         i18 : Int;
         i19 : Int;
         i20 : Int;
         i21 : Int;
      END_STRUCT;
      STC_tMngSysReg : Struct   // Managment system register
         tST : Struct
            xWrite_Request : Bool;
            xDone : Bool;
            xBusy : Bool;
            xError : Bool;
            xSpare4 : Bool;
            xSpare5 : Bool;
            xSpare6 : Bool;
            xSpare7 : Bool;
            ID : Hw_Io;
            dINDEX : DInt;
            uiLEN : UInt;
            dwSTATUS : DWord;
            iSpare : Int;
         END_STRUCT;
         tDATA : Struct
            wRequest_refere_RequestID : Word := W#16#102;   // (Request_referece=01 Alwais=01 )*(RequestID=02 Change Param)
            wAxis_NoOfParameters : Word := W#16#101;   // (Axis=Num.Object)(NoOfParameters=Num of parameter to change)
            wAttribute_NoOfElements : Word := W#16#1001;   // (Attribute=10 Alwais=10)(NoOfParameters=Num of subparameter to Write)
            iParameter_number : Int := 2599;   // Parameter_number=Number of the parameter
            wSubindex : Word;   // Subindex
            wFormat_NoOfValue : Word := W#16#4301;   // (Format_NoOfValue=Format 42=Word 43=Dword)(Num. of value to transfer)
            dwRegisterValue : DWord := DW#16#1;   // Register value
         END_STRUCT;
      END_STRUCT;
      STC_tWriteRecord : WRREC;
      STC_tPZD_OpCLLoop : Struct   // Motor module open/close loop telegram 1
         tR : Struct   // READ
            tZSW1 : Struct   // R2089[0].STATUS WORD 1
               x8 : Bool;   // Speed setp-act val deviation in tollerance
               x9 : Bool;   // Control request
               x10 : Bool;   // F or n comparision value reached or exceeded
               x11 : Bool;   // Tourque limit reached
               x12 : Bool;   // Open holding brake
               x13 : Bool;   // Alarm motor overtemperature
               x14 : Bool;   // n_act>=0
               x15 : Bool;   // Alarm power unit thermal overload
               x0 : Bool;   // Ready for switch on
               x1 : Bool;   // Ready
               x2 : Bool;   // Operation enabled
               x3 : Bool;   // Fault present
               x4 : Bool;   // OFF2
               x5 : Bool;   // OFF3
               x6 : Bool;   // Switching on inhibited active
               x7 : Bool;   // Alarm present
            END_STRUCT;
            iNIST_A : Int;   // R63.Actual speed value
            iFAULT_CODE : Int;   // R2131.Actual fault code
            iWARN_CODE : Int;   // R2132.Actual alarm code
            iUserData1 : Int;
            iUserData2 : Int;
         END_STRUCT;
         tW : Struct   // WRITE
            tSTW1 : Struct   // CONTROL WORD 1
               x8 : Bool;   // Reserved
               x9 : Bool;   // P1122[0].Bypass ramp-function generator
               x10 : Bool;   // P854[0].Control by PLC
               x11 : Bool;   // P1113[0].Setpoint inversion
               x12 : Bool;   // Reserved
               x13 : Bool;   // P1035[0].Motorized potentiometer setpoint raise
               x14 : Bool;   // P1036[0].Motorized potentiometer setpoint lower
               x15 : Bool;   // P855[0] Brake release
               x0 : Bool;   // P840[0].ON/OFF
               x1 : Bool;   // P844[0].OFF2
               x2 : Bool;   // P848[0].OFF3
               x3 : Bool;   // P852[0].Enable operation
               x4 : Bool;   // P1140[0].Enable ramp function generator
               x5 : Bool;   // P1141[0].Continue ramp function generator
               x6 : Bool;   // P1142[0].Enable setpoint
               x7 : Bool;   // P2103[0].Acknowledge faults
            END_STRUCT;
            iNSOLL_A : Int;   // P1070[0].Main set point
            iACC : Int;   // P1138[0].Acceleration ramp % [0-16384]
            iDEC : Int;   // P1139[0].Deceleration ramp % [0-16384]
            iExtRef : Int;   // P1076[0].External reference scaling % [0-16384]
            iUserData2 : Int;
         END_STRUCT;
      END_STRUCT;
   END_VAR
   VAR_TEMP
      TMP_dOldValue_AR1 : DInt;
      TMP_dOldValue_AR2 : DInt;
      TMP_x : Bool;
      TMP_i : Int;
      TMP_d : DInt;
      TMP_r : Real;
      TMP_a : ANY;
      TMP_dZero : DInt;
      TMP_xAlwaysON : Bool;
      TMP_rActualSpeed : Real;
      TMP_iAddressLength : Int;
      TMP_dActualPosMin_dmm : DInt;   // Actual position minimum tollerance [mm/10]
      TMP_dActualPosMax_dmm : DInt;   // Actual position maximum tollerance [mm/10]
      TMP_iRetVal : Int;
   END_VAR
BEGIN

REGION Network 1 (STL): Save AR1 & AR2 value
   //    TAR1
   //    T     #TMP_dOldValue_AR1
   //    TAR2
   //    T     #TMP_dOldValue_AR2
END_REGION

REGION Network 2: #####_COSTANTS_#####
END_REGION

REGION Network 3 (STL): Initializing
         SET;
         S     #TMP_xAlwaysON;

         L     DINT#0;
         T     #TMP_dZero;


         CALL  FILL
         ( BVAL    := #TMP_dZero,
           RET_VAL := #TMP_iRetVal,
           BLK     := #STC_tPZD_OpCLLoop.tR
         );

         CALL  FILL
         ( BVAL    := #TMP_dZero,
           RET_VAL := #TMP_iRetVal,
           BLK     := #STC_tMngSysReg
         );
END_REGION

REGION Network 4: #####_MOTOR_MODULE_#####
END_REGION

REGION Network 5 (STL): Check system data coerence
         L     #STC_tSYS_DATA.iIOAddress_MM;
         L     0;
         <I;
         L     10;
         JC    Err;

         L     #STC_tSYS_DATA.dMaxSpeed_rpm;
         L     DINT#0;
         <=D;
         L     11;
         JC    Err;

         L     #STC_tSYS_DATA.rK_rpm_mmMin;
         L     0.0;
         <=R;
         L     12;
         JC    Err;

         L     #STC_tSYS_DATA.rK_mmMin_Rpm;
         L     0.0;
         <=R;
         L     13;
         JC    Err;

         L     #STC_tSYS_DATA.rMaxAcc_s;
         L     0.0;
         <=R;
         L     14;
         JC    Err;

         L     #STC_tSYS_DATA.rMaxDec_s;
         L     0.0;
         <=R;
         L     15;
         JC    Err;

         L     6;
         T     #TMP_iAddressLength;

   //Compute destination position
         L;
         LAR1;
   //byte 1 = 10h (FIXED for S7)
         L     B#16#10;
         T     B[AR1, P#0.0];
   //byte 2 = data type
         L     B#16#4;  //4 = word
         T     B[AR1, P#1.0];
   //byte 3 & 4 = number of element
         L     #TMP_iAddressLength;  //Production data
         T     W[AR1, P#2.0];
   //byte 5 & 6 = number of DB
         L     0;  //DB production data
         T     W[AR1, P#4.0];
   //byte 7 = memory area
         L     B#16#81;  //81h = I (Input)
         T     B[AR1, P#6.0];
   //byte 8 & 9 = address. Bit 0,1,2 of tenth byte is bit offset
   //byte 7 = address (high). Valid value = 0-7. Bit 3,4,5,6,7 always 0

         L     #STC_tSYS_DATA.iIOAddress_MM;  //Item size
         SLW   3;
         T     W[AR1, P#8.0];
         SRD   16;
         AW    16#0007;
         T     B[AR1, P#7.0];
END_REGION

REGION Network 6: ########################_OPEN_CLOSE_LOOP_#######################
END_REGION

REGION Network 7: #####_MATCH_#####
END_REGION

REGION Network 8 (STL): Input copy
         CALL  BLKMOV
         ( SRCBLK  := #TMP_a,
           RET_VAL := #TMP_iRetVal,
           DSTBLK  := #STC_tPZD_OpCLLoop.tR
         );
END_REGION

REGION Network 9: Status signals
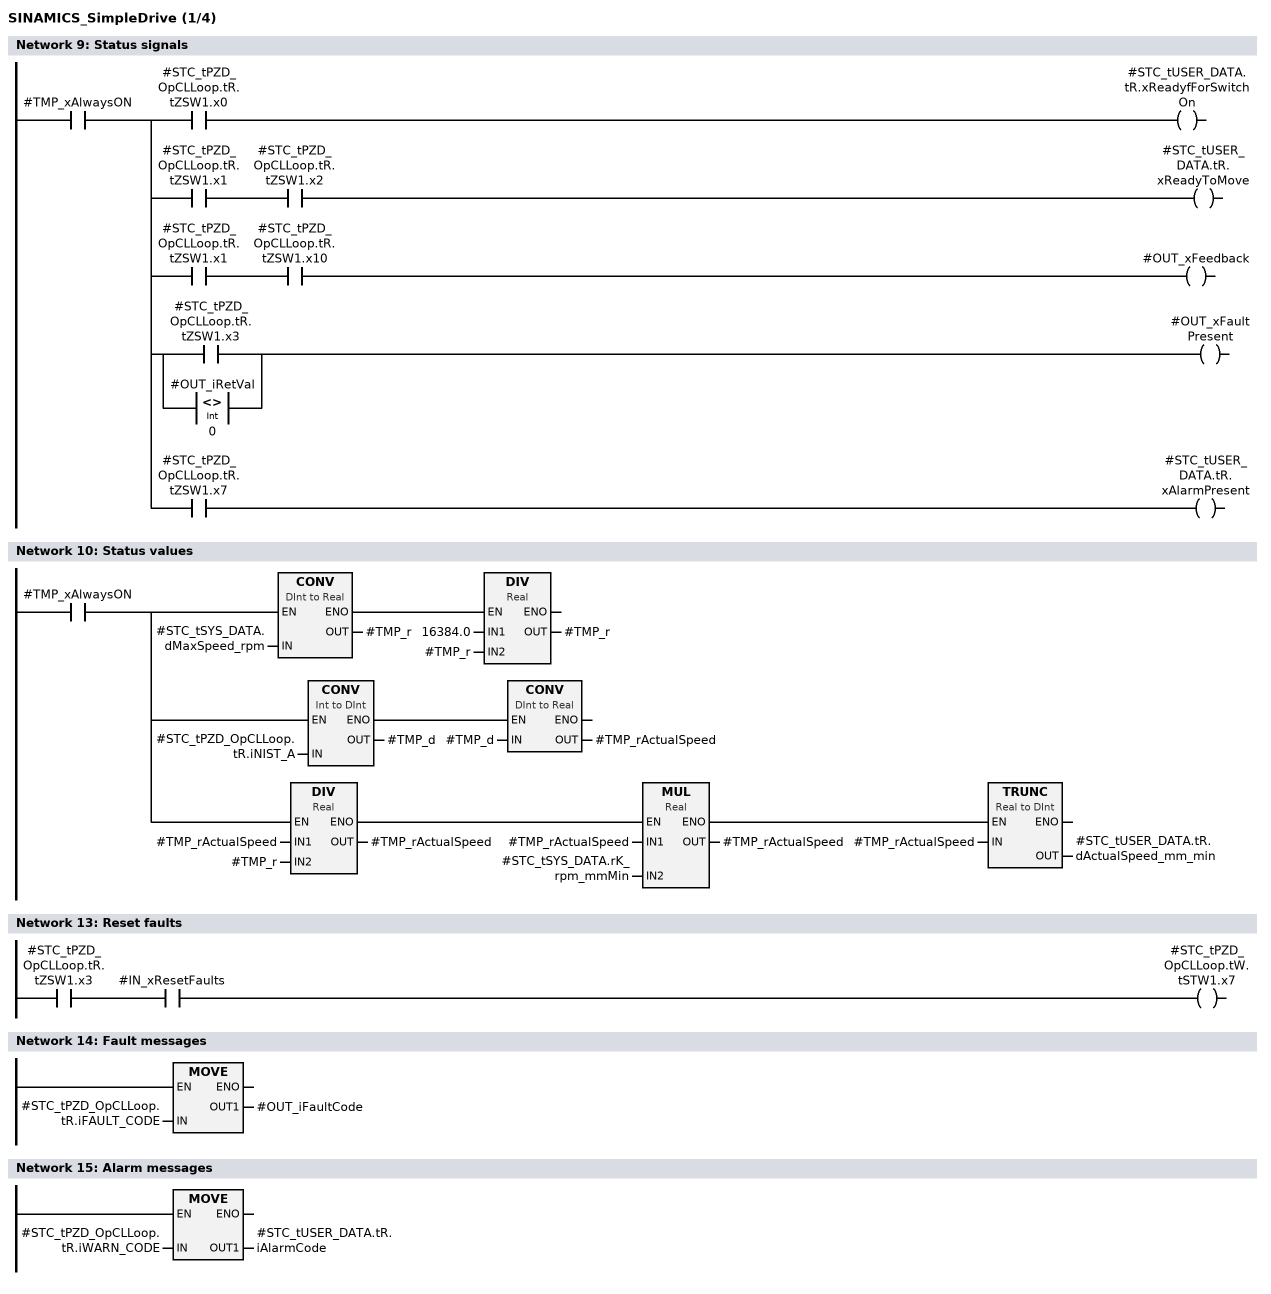
   RUNG wire#powerrail
      Contact( #TMP_xAlwaysON )
      wire#w1
      Contact( #STC_tPZD_OpCLLoop.tR.tZSW1.x0 )
      Coil( #STC_tUSER_DATA.tR.xReadyfForSwitchOn )
   END_RUNG
   RUNG wire#w1
      Contact( #STC_tPZD_OpCLLoop.tR.tZSW1.x1 )
      Contact( #STC_tPZD_OpCLLoop.tR.tZSW1.x2 )
      Coil( #STC_tUSER_DATA.tR.xReadyToMove )
   END_RUNG
   RUNG wire#w1
      Contact( #STC_tPZD_OpCLLoop.tR.tZSW1.x1 )
      Contact( #STC_tPZD_OpCLLoop.tR.tZSW1.x10 )
      Coil( #OUT_xFeedback )
   END_RUNG
   RUNG wire#w1
      Contact( #STC_tPZD_OpCLLoop.tR.tZSW1.x3 )
      wire#w2
      Coil( #OUT_xFaultPresent )
   END_RUNG
   RUNG wire#w1
      { S7_Templates := "SrcType := Int" } NE_Contact(in1 := #OUT_iRetVal, in2 := 0)
   END_RUNG wire#w2
   RUNG wire#w1
      Contact( #STC_tPZD_OpCLLoop.tR.tZSW1.x7 )
      Coil( #STC_tUSER_DATA.tR.xAlarmPresent )
   END_RUNG
   // the same network as SCL:
   #STC_tUSER_DATA.tR.xReadyfForSwitchOn := #TMP_xAlwaysON AND #STC_tPZD_OpCLLoop.tR.tZSW1.x0;
   #STC_tUSER_DATA.tR.xReadyToMove := #TMP_xAlwaysON AND #STC_tPZD_OpCLLoop.tR.tZSW1.x1 AND #STC_tPZD_OpCLLoop.tR.tZSW1.x2;
   #OUT_xFeedback := #TMP_xAlwaysON AND #STC_tPZD_OpCLLoop.tR.tZSW1.x1 AND #STC_tPZD_OpCLLoop.tR.tZSW1.x10;
   #OUT_xFaultPresent := #TMP_xAlwaysON AND (#STC_tPZD_OpCLLoop.tR.tZSW1.x3 OR (#OUT_iRetVal <> 0));
   #STC_tUSER_DATA.tR.xAlarmPresent := #TMP_xAlwaysON AND #STC_tPZD_OpCLLoop.tR.tZSW1.x7;
END_REGION

REGION Network 10: Status values
   RUNG wire#powerrail
      Contact( #TMP_xAlwaysON )
      wire#w1
      { S7_Templates := "[SrcType := DInt, DestType := Real]"; S7_GenerateENO := "TRUE" } Convert(in := #STC_tSYS_DATA.dMaxSpeed_rpm, out => #TMP_r)
      { S7_Templates := "SrcType := Real"; S7_GenerateENO := "TRUE" } Div(in1 := 16384.0, in2 := #TMP_r, out => #TMP_r)
   END_RUNG
   RUNG wire#w1
      { S7_Templates := "[SrcType := Int, DestType := DInt]"; S7_GenerateENO := "TRUE" } Convert(in := #STC_tPZD_OpCLLoop.tR.iNIST_A, out => #TMP_d)
      { S7_Templates := "[SrcType := DInt, DestType := Real]"; S7_GenerateENO := "TRUE" } Convert(in := #TMP_d, out => #TMP_rActualSpeed)
   END_RUNG
   RUNG wire#w1
      { S7_Templates := "SrcType := Real"; S7_GenerateENO := "TRUE" } Div(in1 := #TMP_rActualSpeed, in2 := #TMP_r, out => #TMP_rActualSpeed)
      { S7_Templates := "SrcType := Real"; S7_GenerateENO := "TRUE" } Mul(in1 := #TMP_rActualSpeed, in2 := #STC_tSYS_DATA.rK_rpm_mmMin, out => #TMP_rActualSpeed)
      { S7_Templates := "[SrcType := Real, DestType := DInt]"; S7_GenerateENO := "TRUE" } Trunc(in := #TMP_rActualSpeed, out => #STC_tUSER_DATA.tR.dActualSpeed_mm_min)
   END_RUNG
   // the same network as SCL:
   // ENO of a box is taken as its EN; it also drops when the box reports an error
   IF #TMP_xAlwaysON THEN
       #TMP_r := DINT_TO_REAL(#STC_tSYS_DATA.dMaxSpeed_rpm);
       #TMP_r := 16384.0 / #TMP_r;
       #TMP_d := INT_TO_DINT(#STC_tPZD_OpCLLoop.tR.iNIST_A);
       #TMP_rActualSpeed := DINT_TO_REAL(#TMP_d);
       #TMP_rActualSpeed := #TMP_rActualSpeed / #TMP_r;
       #TMP_rActualSpeed := #TMP_rActualSpeed * #STC_tSYS_DATA.rK_rpm_mmMin;
       #STC_tUSER_DATA.tR.dActualSpeed_mm_min := TRUNC(#TMP_rActualSpeed);
   END_IF;
END_REGION

REGION Network 11: #####_STATUSES_#####
END_REGION

REGION Network 12: #####_ALARMS_#####
END_REGION

REGION Network 13: Reset faults
   RUNG wire#powerrail
      Contact( #STC_tPZD_OpCLLoop.tR.tZSW1.x3 )
      Contact( #IN_xResetFaults )
      Coil( #STC_tPZD_OpCLLoop.tW.tSTW1.x7 )
   END_RUNG
   // the same network as SCL:
   #STC_tPZD_OpCLLoop.tW.tSTW1.x7 := #STC_tPZD_OpCLLoop.tR.tZSW1.x3 AND #IN_xResetFaults;
END_REGION

REGION Network 14: Fault messages
   RUNG wire#powerrail
      { S7_GenerateENO := "TRUE" } Move(in := #STC_tPZD_OpCLLoop.tR.iFAULT_CODE, out1 => #OUT_iFaultCode)
   END_RUNG
   // the same network as SCL:
   #OUT_iFaultCode := #STC_tPZD_OpCLLoop.tR.iFAULT_CODE;
END_REGION

REGION Network 15: Alarm messages
   RUNG wire#powerrail
      { S7_GenerateENO := "TRUE" } Move(in := #STC_tPZD_OpCLLoop.tR.iWARN_CODE, out1 => #STC_tUSER_DATA.tR.iAlarmCode)
   END_RUNG
   // the same network as SCL:
   #STC_tUSER_DATA.tR.iAlarmCode := #STC_tPZD_OpCLLoop.tR.iWARN_CODE;
END_REGION

REGION Network 16: #####_PHASES_&_LOGICS_#####
END_REGION

REGION Network 17: Enable PLC control
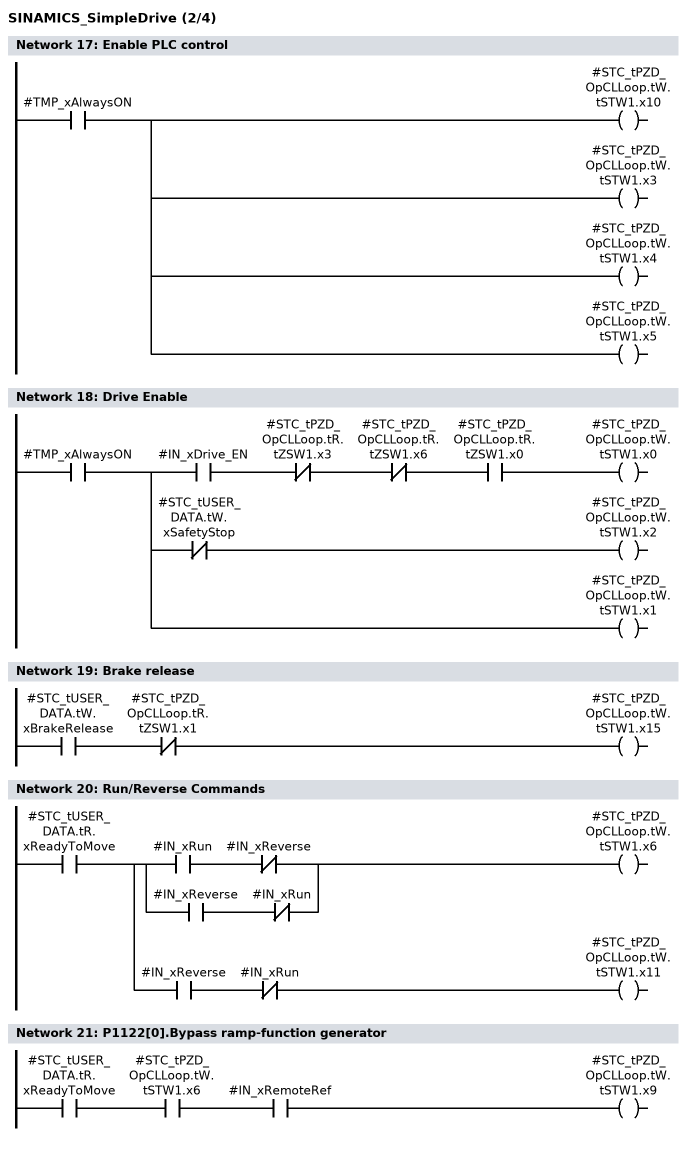
   RUNG wire#powerrail
      Contact( #TMP_xAlwaysON )
      wire#w1
      Coil( #STC_tPZD_OpCLLoop.tW.tSTW1.x10 )
   END_RUNG
   RUNG wire#w1
      Coil( #STC_tPZD_OpCLLoop.tW.tSTW1.x3 )
   END_RUNG
   RUNG wire#w1
      Coil( #STC_tPZD_OpCLLoop.tW.tSTW1.x4 )
   END_RUNG
   RUNG wire#w1
      Coil( #STC_tPZD_OpCLLoop.tW.tSTW1.x5 )
   END_RUNG
   // the same network as SCL:
   #STC_tPZD_OpCLLoop.tW.tSTW1.x10 := #TMP_xAlwaysON;
   #STC_tPZD_OpCLLoop.tW.tSTW1.x3 := #TMP_xAlwaysON;
   #STC_tPZD_OpCLLoop.tW.tSTW1.x4 := #TMP_xAlwaysON;
   #STC_tPZD_OpCLLoop.tW.tSTW1.x5 := #TMP_xAlwaysON;
END_REGION

REGION Network 18: Drive Enable
   RUNG wire#powerrail
      Contact( #TMP_xAlwaysON )
      wire#w1
      Contact( #IN_xDrive_EN )
      I_Contact( #STC_tPZD_OpCLLoop.tR.tZSW1.x3 )
      I_Contact( #STC_tPZD_OpCLLoop.tR.tZSW1.x6 )
      Contact( #STC_tPZD_OpCLLoop.tR.tZSW1.x0 )
      Coil( #STC_tPZD_OpCLLoop.tW.tSTW1.x0 )
   END_RUNG
   RUNG wire#w1
      I_Contact( #STC_tUSER_DATA.tW.xSafetyStop )
      Coil( #STC_tPZD_OpCLLoop.tW.tSTW1.x2 )
   END_RUNG
   RUNG wire#w1
      Coil( #STC_tPZD_OpCLLoop.tW.tSTW1.x1 )
   END_RUNG
   // the same network as SCL:
   #STC_tPZD_OpCLLoop.tW.tSTW1.x0 := #TMP_xAlwaysON AND #IN_xDrive_EN AND NOT #STC_tPZD_OpCLLoop.tR.tZSW1.x3 AND NOT #STC_tPZD_OpCLLoop.tR.tZSW1.x6 AND #STC_tPZD_OpCLLoop.tR.tZSW1.x0;
   #STC_tPZD_OpCLLoop.tW.tSTW1.x2 := #TMP_xAlwaysON AND NOT #STC_tUSER_DATA.tW.xSafetyStop;
   #STC_tPZD_OpCLLoop.tW.tSTW1.x1 := #TMP_xAlwaysON;
END_REGION

REGION Network 19: Brake release
   RUNG wire#powerrail
      Contact( #STC_tUSER_DATA.tW.xBrakeRelease )
      I_Contact( #STC_tPZD_OpCLLoop.tR.tZSW1.x1 )
      Coil( #STC_tPZD_OpCLLoop.tW.tSTW1.x15 )
   END_RUNG
   // the same network as SCL:
   #STC_tPZD_OpCLLoop.tW.tSTW1.x15 := #STC_tUSER_DATA.tW.xBrakeRelease AND NOT #STC_tPZD_OpCLLoop.tR.tZSW1.x1;
END_REGION

REGION Network 20: Run/Reverse Commands
   RUNG wire#powerrail
      Contact( #STC_tUSER_DATA.tR.xReadyToMove )
      wire#w1
      Contact( #IN_xRun )
      I_Contact( #IN_xReverse )
      wire#w2
      Coil( #STC_tPZD_OpCLLoop.tW.tSTW1.x6 )
   END_RUNG
   RUNG wire#w1
      Contact( #IN_xReverse )
      I_Contact( #IN_xRun )
   END_RUNG wire#w2
   RUNG wire#w1
      Contact( #IN_xReverse )
      I_Contact( #IN_xRun )
      Coil( #STC_tPZD_OpCLLoop.tW.tSTW1.x11 )
   END_RUNG
   // the same network as SCL:
   #STC_tPZD_OpCLLoop.tW.tSTW1.x6 := #STC_tUSER_DATA.tR.xReadyToMove AND ((#IN_xRun AND NOT #IN_xReverse) OR (#IN_xReverse AND NOT #IN_xRun));
   #STC_tPZD_OpCLLoop.tW.tSTW1.x11 := #STC_tUSER_DATA.tR.xReadyToMove AND #IN_xReverse AND NOT #IN_xRun;
END_REGION

REGION Network 21: P1122[0].Bypass ramp-function generator
   RUNG wire#powerrail
      Contact( #STC_tUSER_DATA.tR.xReadyToMove )
      Contact( #STC_tPZD_OpCLLoop.tW.tSTW1.x6 )
      Contact( #IN_xRemoteRef )
      Coil( #STC_tPZD_OpCLLoop.tW.tSTW1.x9 )
   END_RUNG
   // the same network as SCL:
   #STC_tPZD_OpCLLoop.tW.tSTW1.x9 := #STC_tUSER_DATA.tR.xReadyToMove AND #STC_tPZD_OpCLLoop.tW.tSTW1.x6 AND #IN_xRemoteRef;
END_REGION

REGION Network 22: #####_PARAMETERS_#####
END_REGION

REGION Network 23: Speed
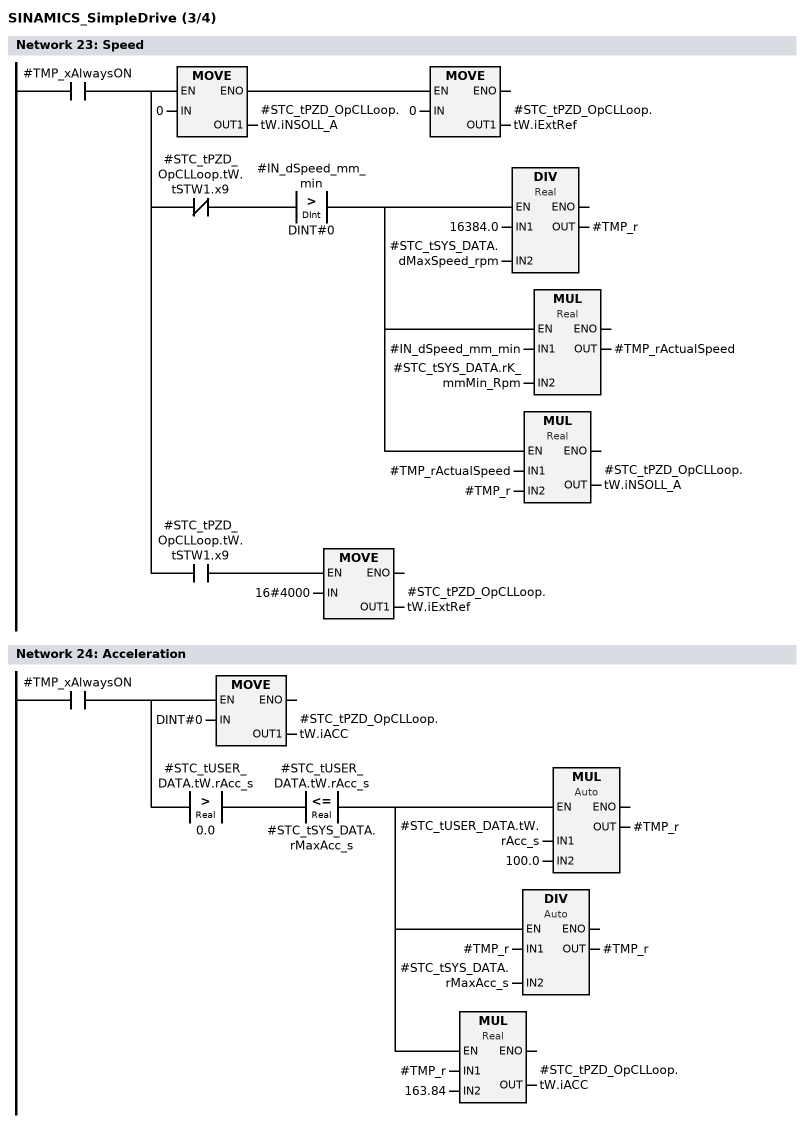
   RUNG wire#powerrail
      Contact( #TMP_xAlwaysON )
      wire#w1
      Move(in := 0, out1 => #STC_tPZD_OpCLLoop.tW.iNSOLL_A)
      Move(in := 0, out1 => #STC_tPZD_OpCLLoop.tW.iExtRef)
   END_RUNG
   RUNG wire#w1
      I_Contact( #STC_tPZD_OpCLLoop.tW.tSTW1.x9 )
      { S7_Templates := "SrcType := DInt" } GT_Contact(in1 := #IN_dSpeed_mm_min, in2 := DINT#0)
      wire#w2
      { S7_Templates := "SrcType := Real" } Div(in1 := 16384.0, in2 := #STC_tSYS_DATA.dMaxSpeed_rpm, out => #TMP_r)
   END_RUNG
   RUNG wire#w2
      { S7_Templates := "SrcType := Real" } Mul(in1 := #IN_dSpeed_mm_min, in2 := #STC_tSYS_DATA.rK_mmMin_Rpm, out => #TMP_rActualSpeed)
   END_RUNG
   RUNG wire#w2
      { S7_Templates := "SrcType := Real" } Mul(in1 := #TMP_rActualSpeed, in2 := #TMP_r, out => #STC_tPZD_OpCLLoop.tW.iNSOLL_A)
   END_RUNG
   RUNG wire#w1
      Contact( #STC_tPZD_OpCLLoop.tW.tSTW1.x9 )
      Move(in := 16#4000, out1 => #STC_tPZD_OpCLLoop.tW.iExtRef)
   END_RUNG
   // the same network as SCL:
   IF #TMP_xAlwaysON THEN
       #STC_tPZD_OpCLLoop.tW.iNSOLL_A := 0;
       #STC_tPZD_OpCLLoop.tW.iExtRef := 0;
   END_IF;
   IF #TMP_xAlwaysON AND NOT #STC_tPZD_OpCLLoop.tW.tSTW1.x9 AND (#IN_dSpeed_mm_min > DINT#0) THEN
       #TMP_r := 16384.0 / #STC_tSYS_DATA.dMaxSpeed_rpm;
       #TMP_rActualSpeed := #IN_dSpeed_mm_min * #STC_tSYS_DATA.rK_mmMin_Rpm;
       #STC_tPZD_OpCLLoop.tW.iNSOLL_A := #TMP_rActualSpeed * #TMP_r;
   END_IF;
   IF #TMP_xAlwaysON AND #STC_tPZD_OpCLLoop.tW.tSTW1.x9 THEN
       #STC_tPZD_OpCLLoop.tW.iExtRef := 16#4000;
   END_IF;
END_REGION

REGION Network 24: Acceleration
   RUNG wire#powerrail
      Contact( #TMP_xAlwaysON )
      wire#w1
      Move(in := DINT#0, out1 => #STC_tPZD_OpCLLoop.tW.iACC)
   END_RUNG
   RUNG wire#w1
      { S7_Templates := "SrcType := Real" } GT_Contact(in1 := #STC_tUSER_DATA.tW.rAcc_s, in2 := 0.0)
      { S7_Templates := "SrcType := Real" } LE_Contact(in1 := #STC_tUSER_DATA.tW.rAcc_s, in2 := #STC_tSYS_DATA.rMaxAcc_s)
      wire#w2
      Mul(in1 := #STC_tUSER_DATA.tW.rAcc_s, in2 := 100.0, out => #TMP_r)
   END_RUNG
   RUNG wire#w2
      Div(in1 := #TMP_r, in2 := #STC_tSYS_DATA.rMaxAcc_s, out => #TMP_r)
   END_RUNG
   RUNG wire#w2
      { S7_Templates := "SrcType := Real" } Mul(in1 := #TMP_r, in2 := 163.84, out => #STC_tPZD_OpCLLoop.tW.iACC)
   END_RUNG
   // the same network as SCL:
   IF #TMP_xAlwaysON THEN #STC_tPZD_OpCLLoop.tW.iACC := DINT#0; END_IF;
   IF #TMP_xAlwaysON AND (#STC_tUSER_DATA.tW.rAcc_s > 0.0) AND (#STC_tUSER_DATA.tW.rAcc_s <= #STC_tSYS_DATA.rMaxAcc_s) THEN
       #TMP_r := #STC_tUSER_DATA.tW.rAcc_s * 100.0;
       #TMP_r := #TMP_r / #STC_tSYS_DATA.rMaxAcc_s;
       #STC_tPZD_OpCLLoop.tW.iACC := #TMP_r * 163.84;
   END_IF;
END_REGION

REGION Network 25: Deceleration
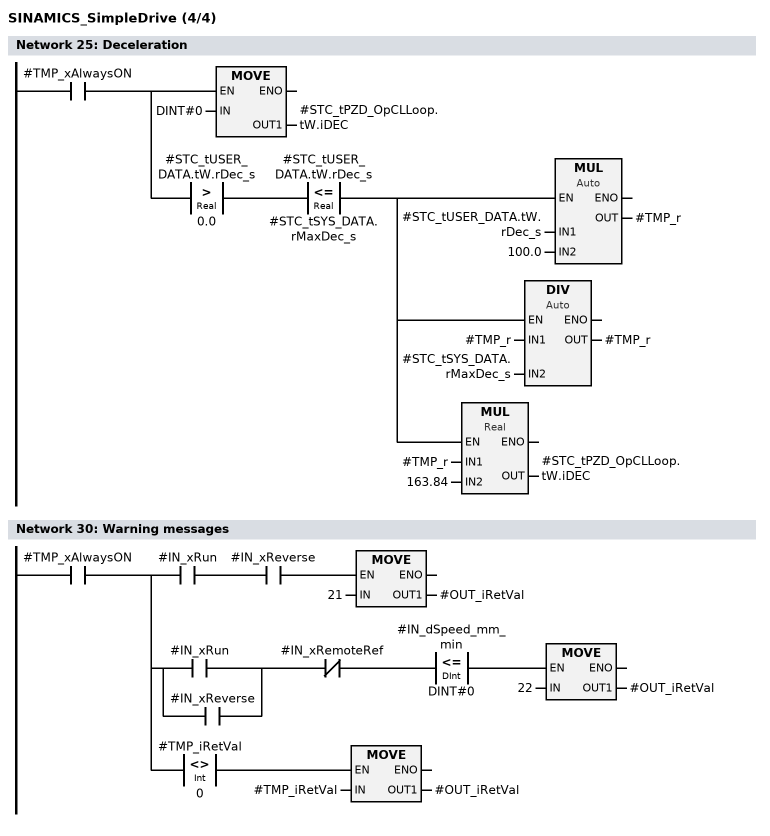
   RUNG wire#powerrail
      Contact( #TMP_xAlwaysON )
      wire#w1
      Move(in := DINT#0, out1 => #STC_tPZD_OpCLLoop.tW.iDEC)
   END_RUNG
   RUNG wire#w1
      { S7_Templates := "SrcType := Real" } GT_Contact(in1 := #STC_tUSER_DATA.tW.rDec_s, in2 := 0.0)
      { S7_Templates := "SrcType := Real" } LE_Contact(in1 := #STC_tUSER_DATA.tW.rDec_s, in2 := #STC_tSYS_DATA.rMaxDec_s)
      wire#w2
      Mul(in1 := #STC_tUSER_DATA.tW.rDec_s, in2 := 100.0, out => #TMP_r)
   END_RUNG
   RUNG wire#w2
      Div(in1 := #TMP_r, in2 := #STC_tSYS_DATA.rMaxDec_s, out => #TMP_r)
   END_RUNG
   RUNG wire#w2
      { S7_Templates := "SrcType := Real" } Mul(in1 := #TMP_r, in2 := 163.84, out => #STC_tPZD_OpCLLoop.tW.iDEC)
   END_RUNG
   // the same network as SCL:
   IF #TMP_xAlwaysON THEN #STC_tPZD_OpCLLoop.tW.iDEC := DINT#0; END_IF;
   IF #TMP_xAlwaysON AND (#STC_tUSER_DATA.tW.rDec_s > 0.0) AND (#STC_tUSER_DATA.tW.rDec_s <= #STC_tSYS_DATA.rMaxDec_s) THEN
       #TMP_r := #STC_tUSER_DATA.tW.rDec_s * 100.0;
       #TMP_r := #TMP_r / #STC_tSYS_DATA.rMaxDec_s;
       #STC_tPZD_OpCLLoop.tW.iDEC := #TMP_r * 163.84;
   END_IF;
END_REGION

REGION Network 26: ################_MOTOR_MODULE_TELEGRAMS_ENDING_#################
END_REGION

REGION Network 27 (STL): Output copy motor module
         L     6;
         T     #TMP_iAddressLength;

   //Compute destination position
         L;
         LAR1;
   //byte 1 = 10h (FIXED for S7)
         L     B#16#10;
         T     B[AR1, P#0.0];
   //byte 2 = data type
         L     B#16#4;  //4 = word
         T     B[AR1, P#1.0];
   //byte 3 & 4 = number of element
         L     #TMP_iAddressLength;  //Production data
         T     W[AR1, P#2.0];
   //byte 5 & 6 = number of DB
         L     0;  //DB production data
         T     W[AR1, P#4.0];
   //byte 7 = memory area
         L     B#16#82;  //82h = Q (Output)
         T     B[AR1, P#6.0];
   //byte 8 & 9 = address. Bit 0,1,2 of tenth byte is bit offset
   //byte 7 = address (high). Valid value = 0-7. Bit 3,4,5,6,7 always 0
         L     #STC_tSYS_DATA.iIOAddress_MM;  //Item size
         SLW   3;
         T     W[AR1, P#8.0];
         SRD   16;
         AW    16#0007;
         T     B[AR1, P#7.0];

         CALL  BLKMOV
         ( SRCBLK  := #STC_tPZD_OpCLLoop.tW,
           RET_VAL := #TMP_iRetVal,
           DSTBLK  := #TMP_a
         );
END_REGION

REGION Network 28: #####_RETVAL_RESPONSE_#####
END_REGION

REGION Network 29 (STL): Initialize RetVal
         L     0;
         T     #OUT_iRetVal;
END_REGION

REGION Network 30: Warning messages
   RUNG wire#powerrail
      Contact( #TMP_xAlwaysON )
      wire#w1
      Contact( #IN_xRun )
      Contact( #IN_xReverse )
      { S7_GenerateENO := "TRUE" } Move(in := 21, out1 => #OUT_iRetVal)
   END_RUNG
   RUNG wire#w1
      Contact( #IN_xRun )
      wire#w2
      I_Contact( #IN_xRemoteRef )
      { S7_Templates := "SrcType := DInt" } LE_Contact(in1 := #IN_dSpeed_mm_min, in2 := DINT#0)
      { S7_GenerateENO := "TRUE" } Move(in := 22, out1 => #OUT_iRetVal)
   END_RUNG
   RUNG wire#w1
      Contact( #IN_xReverse )
   END_RUNG wire#w2
   RUNG wire#w1
      { S7_Templates := "SrcType := Int" } NE_Contact(in1 := #TMP_iRetVal, in2 := 0)
      { S7_GenerateENO := "TRUE" } Move(in := #TMP_iRetVal, out1 => #OUT_iRetVal)
   END_RUNG
   // the same network as SCL:
   IF #TMP_xAlwaysON AND #IN_xRun AND #IN_xReverse THEN #OUT_iRetVal := 21; END_IF;
   IF #TMP_xAlwaysON AND (#IN_xRun OR #IN_xReverse) AND NOT #IN_xRemoteRef AND (#IN_dSpeed_mm_min <= DINT#0) THEN
       #OUT_iRetVal := 22;
   END_IF;
   IF #TMP_xAlwaysON AND (#TMP_iRetVal <> 0) THEN #OUT_iRetVal := #TMP_iRetVal; END_IF;
END_REGION

REGION Network 31 (STL): Blocking messages
         JU    Rest;
   Err:  T     #OUT_iRetVal;
END_REGION

REGION Network 32 (STL): Reset input commands
   // R     #USER_DATA.W.SafetyStop
   //       R     #USER_DATA.W.FlyChange
   //       R     #USER_DATA.W.PH_Select
   //       R     #USER_DATA.W.StartCountOnHead
   //       R     #USER_DATA.W.StartCountOnTail
   //       R     #USER_DATA.W.BrakeRelease
   //       R     #USER_DATA.W.ResetCount
   //       R     #USER_DATA.W.PresetRq
   //       R     #USER_DATA.W.HomeSearch
   //       R     #USER_DATA.W.ReverseHoming
   //       R     #USER_DATA.W.ReferenceCam
   //       R     #USER_DATA.W.ReferenceZero
   //       R     #USER_DATA.W.MDI_Continue
   //       R     #USER_DATA.W.SwLimitsEnable
   //       R     #USER_DATA.W.HwLimitsEnable
   //       R     #Run
   //       R     #Reverse
   //       R     #RemoteRef
   // 
   //       L     L#0
   //       T     #Speed
   //       T     #USER_DATA.W.Override
   //       T     #USER_DATA.W.Target
   //       T     #USER_DATA.W.Preset
   //       T     #USER_DATA.W.Acc
   //       T     #USER_DATA.W.Dec
   Rest: NOP   0;
   //    SET
   //    R     #IN_xDrive_EN
   //    R     #IN_xResetFaults
END_REGION

REGION Network 33 (STL): Restore AR1 & AR2 value
   //    L     #TMP_dOldValue_AR1
   //    LAR1
   //    L     #TMP_dOldValue_AR2
   //    LAR2
END_REGION
END_FUNCTION_BLOCK

FUNCTION_BLOCK "SINAMICS_LinearPosLT"   // FB54, LAD
TITLE = Sinamics drive manager
{ S7_Optimized_Access := 'FALSE' }
AUTHOR : Armitano
VERSION : 1.4
// Return value:
// * 0: OK
// Blocking message:
// * group 1 to 9: general error
// * group 10 to 19: system data error
//   * 10: Sinamics input/output addresses wrong or not setted
//   * 11: Maximum speed in Rpm wrong or not setted
//   * 12: Conversion coefficent for Rpm/mmMin wrong or not setted
//   * 13: Conversion coefficent for mmMin/Rpm wrong or not setted
//   * 14: Maximum acceleration wrong or not setted
//   * 15: Maximum deceleration wrong or not setted
//   * 19: Comunication telegram numxer unknown
// Warning message:
// * group 20 to 29: user data error
//   * 20: Reference cam signal + reference zero signal no possible
//   * 21: Run command + reverse command no possible
//   * 22: Preset speed at zero during run/reverse command
//   * 23: Run/reverse command during homing command no possible
//   * 24: Absolute positioining no possible without axes referenced
//   * 25: Preset override at zero during run/reverse command
// Other:
// * group 30 to 32: preset data error
//   * 30: Error during send preset value (Check parameters in Sys_Data)
//   * 31: Error during preset command (Check parameters in Sys_Data)
//   * 32: Error during saving preset command (Check Sys_Data)
//   * 34: Error during send preset homing (Check parameters in Sys_Data)
//   * 40: Error during request misured values (Check Sys_Data)
//   * 41: Error during response misured values (Check Sys_Data)
// * group 8000 to 9000: SFC20 code (Read the SFC20 Help)
   VAR_INPUT
      IN_xDrive_EN : Bool;   // Drive enable
      IN_xRun : Bool;   // Run forward
      IN_xReverse : Bool;   // Run backward
      IN_xPositioning : Bool;   // Positioning enable
      IN_xResetFaults : Bool;   // Reset faults
      IN_dSpeed_mm_min : DInt;   // Speed reference [mm/min]
   END_VAR
   VAR_OUTPUT
      OUT_xFeedback : Bool;   // Feedback active
      OUT_xFaultPresent : Bool;   // Fault present
      OUT_iFaultCode : Int;   // Fault code
      OUT_iRetVal : Int;   // Return value in case of wrong configuration
   END_VAR
   VAR
      STC_tUSER_DATA : Struct   // User data (Extended functions commands for execute the application desired)
         tR : Struct
            xReadyfForSwitchOn : Bool;   // Ready for switch on
            xReadyToMove : Bool;   // Ready to move
            xAxleRefered : Bool;   // Axle referenced
            xPositionReached : Bool;   // Position reached
            xAlarmPresent : Bool;   // Alarm present
            xAxleToZero : Bool;   // Axle to zero value
            xAxleAcc : Bool;   // Axle in acceleration
            xAxleDec : Bool;   // Axle in deceleration
            iAlarmCode : Int;   // Alarm code
            dActualPosition_dmm : DInt;   // Actual position value [mm/10]
            dActualSpeed_mm_min : DInt;   // Actual speed value [mm/min]
         END_STRUCT;
         tW : Struct
            xSafetyStop : Bool;   // Safety stop (OFF3)
            xFlyChange : Bool;   // Fly change
            xPH_Select : Bool;   // Photocell selection
            xStartCountOnHead : Bool;   // Start count on glass head
            xStartCountOnTail : Bool;   // Start count on glass tail
            xBrakeRelease : Bool;   // Brake release
            xResetCount : Bool;   // Reset counter
            x8 : Bool;
            x9 : Bool;
            x10 : Bool;
            x11 : Bool;
            x12 : Bool;
            xMDI_Continue : Bool;   // MDI movement continue (only for gearing axes)
            x14 : Bool;
            xHwLimitsEnable : Bool;   // Hardware limits activation
            xEdgePulseStartCount : Bool;   // Edge pulse of start count photocell (for positioning with photocell)
            iOverride_perc : Int := 100;   // Override [%]
            dTarget_dmm : DInt;   // Target position [mm/10]
            d3 : DInt;
            rAcc_m_s2 : Real;   // Acceleration [m/s2]
            rDec_m_s2 : Real;   // Deceleration [m/s2]
         END_STRUCT;
      END_STRUCT;
      STC_tSYS_DATA : Struct   // System data (Info about applications type and HW config.)
         iIOAddress_MM : Int := -1;   // Input/Output addresses for motor module
         i2 : Int;
         i3 : Int;
         i4 : Int;
         i5 : Int;
         i6 : Int;
         i7 : Int;
         dMaxSpeed_rpm : DInt;   // MaxSpeed [rpm]
         d9 : DInt;
         dPosWindow_dmm : DInt := L#1;   // Positioning window [mm/10]
         d11 : DInt;
         d12 : DInt;
         d13 : DInt;
         rK_rpm_mmMin : Real;   // K Conversion from rpm to mm/min
         r15 : Real;
         rMaxAcc_m_s2 : Real;   // MaxAcc [m/s2]
         rMaxDec_m_s2 : Real;   // MaxDec [m/s2]
         r18 : Real;
         r19 : Real;
      END_STRUCT;
      STC_tEXT_DATA : Struct   // Extended data (Functions commands for DCC applications)
         DisGearingCtrl : Bool;   // Disable gearing tollerance error control (Only for gearing axes)
         x1 : Bool;
         x2 : Bool;
         x3 : Bool;
         x4 : Bool;
         ModuleCorrect : Bool;   // Enable module correction (Only positioner with turnover endless)
         x6 : Bool;
         x7 : Bool;
         x8 : Bool;
         x9 : Bool;
         x10 : Bool;
         x11 : Bool;
         x12 : Bool;
         x13 : Bool;
         x14 : Bool;
         x15 : Bool;
         D0 : DInt;
         D1 : DInt;
         D2 : DInt;
         D3 : DInt;
         D4 : DInt;
         D5 : DInt;
         D6 : DInt;
         D7 : DInt;
         D8 : DInt;
         D9 : DInt;
         D10 : DInt;
         D11 : DInt;
      END_STRUCT;
      STC_tST : Struct
         x0 : Bool;   // Positioning Absolute
         x1 : Bool;   // Positioning with photocell
         x2 : Bool;
         x3 : Bool;
         x4 : Bool;
         x5 : Bool;
         x6 : Bool;   // Target = Feedback target
         x7 : Bool;   // Validation position reached with module correction
         x8 : Bool;   // Preset phases in progress
         x9 : Bool;
         x10 : Bool;
         x11 : Bool;   // Axle resetted
         x12 : Bool;
         x13 : Bool;
         x14 : Bool;
         x15 : Bool;
      END_STRUCT;
      STC_tOS_PN : Struct
         x0 : Bool;   // Run
         x1 : Bool;   // Reverse
         x2 : Bool;   // Positioning
         x3 : Bool;   // Fly change
         x4 : Bool;
         x5 : Bool;
         x6 : Bool;   // Waiting photocell signal
         x7 : Bool;   // Position reached
         x8 : Bool;   // Fly referencing active (Positive edge)
         x9 : Bool;   // Fly referencing active (Negative edge)
         x10 : Bool;   // Preset position
         x11 : Bool;
         x12 : Bool;
         x13 : Bool;   // Request misured values
         x14 : Bool;
         x15 : Bool;
      END_STRUCT;
      STC_tOS : Struct
         x0 : Bool;   // Run
         x1 : Bool;   // Reverse
         x2 : Bool;   // Positioning
         x3 : Bool;   // Fly change
         x4 : Bool;
         x5 : Bool;
         x6 : Bool;   // Waiting photocell signal
         x7 : Bool;
         x8 : Bool;   // Fly referencing active
         x9 : Bool;
         x10 : Bool;
         x11 : Bool;
         x12 : Bool;
         x13 : Bool;
         x14 : Bool;
         x15 : Bool;
      END_STRUCT;
      STC_tPH : Struct
         x0 : Bool;   // Positioning initializing
         x1 : Bool;   // Positioning request
         x2 : Bool;   // Fly change waiting
         x3 : Bool;   // Fly change sending
         x4 : Bool;   // Change command waiting
         x5 : Bool;   // Change command request
         x6 : Bool;   // Wait photocell signal
         x7 : Bool;
         x8 : Bool;   // Send encoder value
         x9 : Bool;   // Send preset command
         x10 : Bool;   // Send saving preset command
         x11 : Bool;   // End preset encoder
         x12 : Bool;
         x13 : Bool;   // Request misured values
         x14 : Bool;   // Waiting response values
         x15 : Bool;   // Misured values recived
      END_STRUCT;
      STC_tPROP : Struct
         i0 : Int;   // Previous cycle [ms]
         i1 : Int;
         i2 : Int;   // Override in sending [%]
         d3 : DInt;   // Speed in sending [mm/min]
         d4 : DInt;   // Target in sending [mm/10]
         r5 : Real;   // Acceleration in sending [m/s2]
         r6 : Real;   // Deceleration in sending [m/s2]
         i7 : Int;
         i8 : Int;
         i9 : Int;
         i10 : Int;
         i11 : Int;   // Override in fly change [%]
         d12 : DInt;   // Speed in fly change [mm/min]
         d13 : DInt;   // Target in fly change [mm/10]
         r14 : Real;   // Acceleration in fly change [m/s2]
         r15 : Real;   // Deceleration in fly change [m/s2]
         i16 : Int;
         i17 : Int;
         i18 : Int;
         i19 : Int;
         i20 : Int;
         tmON_feedback_ms : IEC_TIMER;   // Delay feedback [ms]
      END_STRUCT;
      STC_tPZD_Pos : Struct   // Motor module positioner telegram 111
         tR : Struct   // READ
            tZSW1 : Struct   // R2089[0].STATUS WORD 1
               x8 : Bool;   // Tracking error in tolerance
               x9 : Bool;   // Control request
               x10 : Bool;   // Target position reached
               x11 : Bool;   // Reference point set
               x12 : Bool;   // Acknowledgment, traversing block activated
               x13 : Bool;   // In_actl < speed threshold value 3
               x14 : Bool;   // Axis accelerating
               x15 : Bool;   // Axis decelerating
               x0 : Bool;   // Ready for switch on
               x1 : Bool;   // Ready
               x2 : Bool;   // Operation enabled
               x3 : Bool;   // Fault present
               x4 : Bool;   // OFF2
               x5 : Bool;   // OFF3
               x6 : Bool;   // Switching on inhibited active
               x7 : Bool;   // Alarm present
            END_STRUCT;
            tPOS_ZSW1 : Struct   // R2089[3].POSITIONER STATUS WORD 2
               x8 : Bool;   // STOP cam minus active
               x9 : Bool;   // STOP cam plus active
               x10 : Bool;   // Jog active
               x11 : Bool;   // Homing procedure active
               x12 : Bool;   // Flying referencing active
               x13 : Bool;   // Traversing block active
               x14 : Bool;   // Setup active
               x15 : Bool;   // MDI active
               x0 : Bool;   // Active traversing block, bit 0
               x1 : Bool;   // Active traversing block, bit 1
               x2 : Bool;   // Active traversing block, bit 2
               x3 : Bool;   // Active traversing block, bit 3
               x4 : Bool;   // Active traversing block, bit 4
               x5 : Bool;   // Active traversing block, bit 5
               x6 : Bool;   // Reserved
               x7 : Bool;   // Reserved
            END_STRUCT;
            tPOS_ZSW2 : Struct   // R2089[4].POSITIONER STATUS WORD 3
               x8 : Bool;   // Position actual value <= cam switching position 1
               x9 : Bool;   // Position actual value <= cam switching position 2
               x10 : Bool;   // Direct output 1 via traversing block
               x11 : Bool;   // Direct output 2 via traversing block
               x12 : Bool;   // Fixed stop reached
               x13 : Bool;   // Fixed stop clamping torque reached
               x14 : Bool;   // Travel to fixed stop active
               x15 : Bool;   // Traversing command active
               x0 : Bool;   // Tracking mode active
               x1 : Bool;   // Velocity limit active
               x2 : Bool;   // Setpoint available
               x3 : Bool;   // Printing mark outside outer window
               x4 : Bool;   // Axis moves forwards
               x5 : Bool;   // Axis moves backwards
               x6 : Bool;   // Software limit switch minus reached
               x7 : Bool;   // Software limit switch plus reached
            END_STRUCT;
            dFDB_TARGET : DInt;   // R2060[5].Feedback target
            dXIST_A : DInt;   // R2521[0].Actual position value
            dNIST_B : DInt;   // R63.Actual speed value
            iFAULT_CODE : Int;   // R2131.Actual fault code
            iWARN_CODE : Int;   // R2132.Actual alarm code
            iUser : Int;
         END_STRUCT;
         tW : Struct   // WRITE
            tSTW1 : Struct   // CONTROL WORD 1
               x8 : Bool;   // P2589.EPOS jog 1 signal source
               x9 : Bool;   // P2590.EPOS jog 2 signal source
               x10 : Bool;   // P854[0].Control by PLC
               x11 : Bool;   // P2595.EPOS referencing start
               x12 : Bool;   // R2090[12].Enable misure probe
               x13 : Bool;   // P2633.EPOS external block change
               x14 : Bool;   // R2090[14].Disable error tollerance control on gearing axes
               x15 : Bool;   // P855[0].Brake release
               x0 : Bool;   // P840[0].ON/OFF
               x1 : Bool;   // P844[0].OFF2
               x2 : Bool;   // P848[0].OFF3
               x3 : Bool;   // P852[0].Enable operation
               x4 : Bool;   // P2641.EPOS abort traversing task
               x5 : Bool;   // P2640.EPOS intermediate STOP
               x6 : Bool;   // P2631.EPOS activate traversing task
               x7 : Bool;   // P2103.Acknowledge faults
            END_STRUCT;
            tPOS_STW1 : Struct   // POSITIONER CONTROL WORD 2